// TIA Portal project "e045002v093" (V13)

(* hardware
DEVICE "S7-300 station_1"  S7-300 station
   slot 0: "Perfil soporte"  Rail  6ES7 390-1***0-0AA0
   slot 2: "U10.5"  CPU 313C  6ES7 313-5BG04-0AB0  V3.3
      slot 0: "Interfaz MPI_1"  MPI
      slot 2: "DI24/DO16_1"  DI24/DO16
      slot 3: "AI5/AO2_1"  AI5/AO2
      slot 4: "Contaje_1"  Counter
   slot 4: "U7.3"  CP 343-1 LEAN  6GK7 343-1CX10-0XE0  V3.0
   slot 5: "U13.5"  DI32xDC24V  6ES7 321-1BL00-0AA0
   slot 6: "U17.5"  DI32xDC24V  6ES7 321-1BL00-0AA0
   slot 7: "U21.5"  DI32 x 24VDC  6ES7 321-1BL00-0AA0
   slot 8: "U25.5"  DO16xRel. AC120V/230V  6ES7 322-1HH01-0AA0
   slot 9: "U27.5"  DO32xDC24V/0.5A  6ES7 322-1BL00-0AA0
   slot 10: "U35.5"  AO2 x 12bits  6ES7 332-5HB01-0AB0
DEVICE "U9.1"  KTP700 Basic PN
   slot 0: "HMI"  HMI  6AV2 123-2GB03-0AX0  13.0.1.0
   slot 1: "HMI_RT_1"  KTP700 Basic PN  6AV2 123-2GB03-0AX0  13.0.1.0
   slot 5: "U9.1.IE_CP_1"  Interfaz PROFINET
      slot 1: "Interfaz PROFINET_1"  Interfaz PROFINET
         slot 1: "Port_1"  Port
*)

// ===== PLC "U10.5"  CPU 313C =====
// protected blocks, not shown: "FB_CTR_MOT", "FC_MAQ_EST_16", "FC_MAQ_EST_32", "FC_PRC_ALA2", "fbSimContactor"

VAR_GLOBAL   // PLC tag table "00_Tabla de variables estándar"
   "CicIni" AT %M17.2 : Bool;
   "Clock_10.0_Hz" AT %M16.0 : Bool;
   "Clock_5.0_Hz" AT %M16.1 : Bool;
   "Clock_2.5_Hz" AT %M16.2 : Bool;
   "Clock_2.0_Hz" AT %M16.3 : Bool;
   "Clock_1.25_Hz" AT %M16.4 : Bool;
   "Clock_1.0_Hz" AT %M16.5 : Bool;
   "Clock_0.625_Hz" AT %M16.6 : Bool;
   "Clock_0.5_Hz" AT %M16.7 : Bool;
   "bit1" AT %M17.0 : Bool;
   "bit0" AT %M17.1 : Bool;
   "Rec_Todas" AT %M17.3 : Bool;
   "Tag_2" AT %M255.7 : Bool;
   "Tag_3" AT %M255.6 : Bool;
   "Tag_5" AT %M231.0 : Bool;
   "Tag_8" AT %T0 : Timer;
   "Ala_Nue" AT %M17.4 : Bool;
   "Ala_Pre" AT %M17.5 : Bool;
   "Sin_Ala" AT %M17.6 : Bool;
   "Contador" AT %MW18 : Word;
   "xpiSnsAscen_Aba_Par" AT %M248.2 : Bool;
   "_PeticiónPallet" AT %M251.5 : Bool;
   "Tag_9" AT %MB252 : Byte;
   "NoRstFilCompl" AT %M17.7 : Bool;   // No resetear "Fila Completa"
   "Set_TON_iSnsContadEmbal_1" AT %M232.0 : Bool;
   "Tag_4" AT %M241.1 : Bool;
   "Set_TON_iSnsContadEmbal_2" AT %M232.1 : Bool;
   "Set_TON_iSnsPerEmpCajAde" AT %M232.2 : Bool;
   "Cont_iSnsContadEmbal_1" AT %MW100 : Int;
   "Cont_iSnsContadEmbal_2" AT %MW102 : Int;
   "Cont_iSnsPerEmpCajAde" AT %MW104 : Int;
   "Cont_iSnsContadEmbal_3" AT %MW106 : Int;
   "Tag_6" AT %MD110 : Time;
   "Tag_7" AT %MD114 : Time;
   "Tag_10" AT %MD118 : Time;
   "Set_TON_iSnsContadEmbal_3" AT %M232.3 : Bool;
   "Tag_1" AT %T1 : Timer;
   "Tag_11" AT %M254.0 : Bool;
   "Tag_12" AT %M254.1 : Bool;
   "Tag_13" AT %M254.2 : Bool;
   "Tag_14" AT %M254.3 : Bool;
   "Tag_15" AT %M123.5 : Bool;
   "Tag_16" AT %M256.0 : Bool;
   "Tag_1200" AT %M255.0 : Bool;
   "Tag_17" AT %M255.1 : Bool;
   "Tag_18" AT %M33.5 : Bool;
   "Resum_ala_Fech" AT %M33.4 : Bool;
   "Hab_marcha1_2" AT %M50.7 : Bool;
   "T_espera_parada_21.26" AT %M50.5 : Bool;
   "MFRD" AT %M50.4 : Bool;
   "MIGS" AT %M50.6 : Bool;
   "i_SnsFinDosif" AT %I11.0 : Bool;   // Sensor final cinta dosificadora
END_VAR

VAR_GLOBAL   // PLC tag table "240_Memorias_Flancos"
   "xnHMI.Pls_Inc_Elem" AT %M240.0 : Bool;
   "xnHMI.Pls_Dec_Elem" AT %M240.1 : Bool;
   "xnHMI.Pls_Elem_Der" AT %M240.2 : Bool;
   "xnHMI.Pls_Elem_Izq" AT %M240.3 : Bool;
   "xnHMI.Pls_Inc_Fila" AT %M240.4 : Bool;
   "xnHMI.Pls_Dec_Fila" AT %M240.5 : Bool;
   "xnHMI.Pls_Fila_Sup" AT %M240.6 : Bool;
   "xnHMI.Pls_Fila_Inf" AT %M240.7 : Bool;
   "xpHMI.Pls_New_Fila" AT %M241.0 : Bool;
   "xpHMI.Pls_New_Elem" AT %M241.2 : Bool;
   "xpHMI.Pls_Kill_Elem" AT %M241.3 : Bool;
   "xnHMI.Pls_WR_Receta" AT %M241.4 : Bool;
   "xnHMI.Pls_RD_Receta" AT %M241.5 : Bool;
   "xpEditar_Recetas" AT %M241.6 : Bool;
   "xnHMI.Pls_Inc_Receta" AT %M241.7 : Bool;
   "xnHMI.Pls_Dec_Receta" AT %M242.0 : Bool;
   "xnHMI.Pls_Inc_Capa" AT %M242.1 : Bool;
   "xnHMI.Pls_Dec_Capa" AT %M242.2 : Bool;
   "xnHMI.Pls_Elem_+" AT %M242.3 : Bool;
   "xnHMI.Pls_Elem_-" AT %M242.4 : Bool;
   "xpHMI.Pls_CargarReceta" AT %M242.5 : Bool;
   "xpiPul_MarCiclo" AT %M242.6 : Bool;
   "xpiPul_HabTransp" AT %M242.7 : Bool;
   "xpiPul_HabDosif" AT %M243.0 : Bool;
   "xpiPul_HabCargPall" AT %M243.1 : Bool;
   "xpiPul_ResetAla" AT %M243.2 : Bool;
   "xpiSnsContadEmbal_1" AT %M243.3 : Bool;
   "xpiSnsContadEmbal_2" AT %M243.4 : Bool;
   "xniSnsContadEmbal_1" AT %M243.5 : Bool;
   "xniSnsContadEmbal_2" AT %M243.6 : Bool;
   "xpAUTO/MAN" AT %M243.7 : Bool;
   "xnAUTO/MAN" AT %M244.0 : Bool;
   "xniSnsPerEmpCajAde" AT %M244.1 : Bool;
   "xniSnsPallTrnsp_4" AT %M244.2 : Bool;
   "xniSnsPallTrnsp_5" AT %M244.3 : Bool;
   "xpiPul_MultiArr" AT %M244.4 : Bool;
   "xniPul_MultiArr" AT %M244.5 : Bool;
   "xpiPul_MultiAba" AT %M244.6 : Bool;
   "xniPul_MultiAba" AT %M244.7 : Bool;
   "xpiPul_MultiAde" AT %M245.0 : Bool;
   "xniPul_MultiAde" AT %M245.1 : Bool;
   "xpiPul_MultiAtr" AT %M245.2 : Bool;
   "xniPul_MultiAtr" AT %M245.3 : Bool;
   "xpiPul_Multi_A" AT %M245.4 : Bool;
   "xniPul_Multi_A" AT %M245.5 : Bool;
   "xpiPul_Multi_B" AT %M245.6 : Bool;
   "xniPul_Multi_B" AT %M245.7 : Bool;
   "xniSnsPlataf_Ade" AT %M246.0 : Bool;
   "xniSnsPlataf_Atr" AT %M246.1 : Bool;
   "xniSnsPallTrnsp_2" AT %M246.3 : Bool;
   "xpiSnsPallTrnsp_2" AT %M246.2 : Bool;
   "xpiSnsPallRetractil" AT %M246.4 : Bool;
   "xniSnsPallRetractil" AT %M246.5 : Bool;
   "xpiSnsPallTrnsp_4" AT %M246.6 : Bool;
   "xpiSnsPallTrnsp_5" AT %M246.7 : Bool;
   "xpiSnsEmpj_Ade_Par" AT %M247.0 : Bool;
   "xnPALLET_NO_FUERA_ASCENSOR" AT %M247.1 : Bool;
   "xpRECAMBIO_PALLET" AT %M247.2 : Bool;
   "xpiSnsPallEnAscen" AT %M247.3 : Bool;
   "xniSnsPallEnAscen" AT %M247.4 : Bool;
   "xpiSnsAltuPlata_Aba" AT %M247.5 : Bool;
   "xniSnsAltuPlata_Aba" AT %M247.6 : Bool;
   "xpiSnsAltuPlata_Arr" AT %M247.7 : Bool;
   "xniSnsAltuPlata_Arr" AT %M248.0 : Bool;
   "xpiSnsAscen_Arr" AT %M248.1 : Bool;
   "xnEditando_Recetas" AT %M248.3 : Bool;
   "xpHMI.Pls_RD_Receta" AT %M248.4 : Bool;
   "xp3s4" AT %M248.5 : Bool;
   "xp3s9" AT %M248.6 : Bool;
   "xpHMI.Pls_Inc_Figura_Sel" AT %M248.7 : Bool;
   "xpHMI.Pls_Inc_Capa_Editando" AT %M249.0 : Bool;
   "xpHMI.Pls_Dec_Capa_Editando" AT %M249.1 : Bool;
   "xpS_PriElemCapa" AT %M249.2 : Bool;
   "xnElemento_DESCARGADO" AT %M249.3 : Bool;
   "xpiSnsPerEmpCajAde" AT %M249.4 : Bool;
   "xpiSnsContadEmbal_3" AT %M249.5 : Bool;
   "xniSnsContadEmbal_3" AT %M249.6 : Bool;
END_VAR

VAR_GLOBAL   // PLC tag table "20_Recetas"
   "Editando_Recetas" AT %M20.0 : Bool;
   "RECETA_Editando" AT %MB21 : Byte;
   "CAPA_Editando" AT %MB22 : Byte;
END_VAR

VAR_GLOBAL   // PLC tag table "30_Proceso"
   "Elemento_CARGADO" AT %M30.0 : Bool;   // Avanzar en el dibujo
   "Nueva_CAPA" AT %M30.2 : Bool;   // Se terminó una capa
   "Elemento_DESCARGADO" AT %M30.1 : Bool;   // Retroceder en el dibujo
   "Nuevo_PALLET" AT %M30.3 : Bool;   // Se terminó un pallet
   "CICLO_Hab" AT %M30.4 : Bool;   // Máquina en ciclo automático
   "TRANSPORTES_Hab" AT %M30.5 : Bool;
   "DOSIFICADOR_Hab" AT %M30.6 : Bool;
   "CARGAPALLET_Hab" AT %M30.7 : Bool;
   "AUTO/MAN" AT %M31.0 : Bool;   // 1: AUTOMÁTICO / 0: MANUAL
   "ResumAla_Grave" AT %M31.1 : Bool;
   "ResumAla_General" AT %M31.2 : Bool;
   "ResumAla_TranspCaja_1" AT %M31.3 : Bool;
   "ResumAla_TranspCaja_2" AT %M31.4 : Bool;
   "ResumAla_Dosificador_1" AT %M31.5 : Bool;
   "ResumAla_Dosificador_2" AT %M31.6 : Bool;
   "ResumAla_CargaPallet_1" AT %M31.7 : Bool;
   "ResumAla_CargaPallet_2" AT %M32.0 : Bool;
   "ResumAla_CargaPallet_3" AT %M32.1 : Bool;
   "ResumAla_CargaPallet_4" AT %M32.2 : Bool;
   "ResumAla_TranspPall_1" AT %M32.3 : Bool;
   "ResumAla_TranspPall_2" AT %M32.4 : Bool;
   "ResumAla_Warnings" AT %M32.5 : Bool;
   "T_ResumAla_General" AT %M32.6 : Bool;
   "Esperando_Cajas" AT %M32.7 : Bool;
   "Cambio_Elemento" AT %M33.0 : Bool;
   "Elemento_DESCARGADO_scan" AT %M33.1 : Bool;
   "ResumAla_Dosificador_3" AT %M33.2 : Bool;
   "ResumAla_Dosificador_4" AT %M33.3 : Bool;
END_VAR

VAR_GLOBAL   // PLC tag table "Tabla I/O"
   "iPul_MultiArr" AT %E34.0 : Bool;   // Pulsador Multifunción Arriba
   "iPul_MultiAba" AT %E34.1 : Bool;   // Pulsador Multifunción Abajo
   "iPul_MultiAde" AT %E34.2 : Bool;   // Pulsador Multifunción Adelante
   "iPul_MultiAtr" AT %E34.3 : Bool;   // Pulsador Multifunción Atrás
   "iPul_Multi_A" AT %E34.4 : Bool;   // Pulsador Multifunción "A"
   "iPul_Multi_B" AT %E34.5 : Bool;   // Pulsador Multifunción "B"
   "iPul_ResetAla" AT %E34.6 : Bool;   // Pulsador Reset Alarmas
   "iiPul_Emerg" AT %E34.7 : Bool;   // Pulsador Parada de Emergencia en Pupitre
   "iPul_MarCiclo" AT %E32.0 : Bool;   // Pulsador Marcha de Ciclo
   "iiPul_ParaCiclo" AT %E32.1 : Bool;   // Pulsador Parada de Piclo
   "iPul_HabTransp" AT %E32.2 : Bool;   // Pulsador Habilitación Transporte de Entrada
   "iiPul_DeshTransp" AT %E32.3 : Bool;   // Pulsador Deshabilitación Transporte de Entrada
   "iPul_HabDosif" AT %E32.4 : Bool;   // Pulsador Habilitación Dosificador
   "iiPul_DeshDosif" AT %E32.5 : Bool;   // Pulsador Deshabilitación Dosificador
   "iPul_HabCargPall" AT %E32.6 : Bool;   // Pulsador Habilitación Carga de Pallet
   "iiPul_DeshCargPall" AT %E32.7 : Bool;   // Pulsador Deshabilitación Carga de Pallet
   "iSel_Auto/Man" AT %E33.0 : Bool;   // Selectora Automático/Manual
   "iiPul_EmergAlmac_1_AlmacManual" AT %E33.5 : Bool;   // Pulsador Operación Manual Almacén Pallets
   "iiPul_EmergAlmac_2" AT %E1.0 : Bool;   // Pulsador parada de emergencia en almacén
   "iPul_RstSegRetrAlmac" AT %E1.1 : Bool;   // Pulsador reset seguridades retractilador almacén
   "iiPul_EmergAscen" AT %E1.2 : Bool;   // Pulsador parada de emergencia en ascensor
   "iPul_RstSegRetrAscen" AT %E1.3 : Bool;   // Pulsador reset seguridades retractilador ascensor
   "iPul_RstSegRetrEntra" AT %E1.4 : Bool;   // Pulsador reset seguridades retractilador entrada
   "iPul_RstSegRetrSali" AT %E1.5 : Bool;   // Pulsador reset seguridades retractilador salida
   "iiPul_EmergMaq" AT %E1.6 : Bool;   // Pulsador parada de emergencia en máquina
   "iiPul_EmergTransp" AT %E1.7 : Bool;   // Pulsador parada de emergencia en transportes de alimentación
   "iVarEmpj_FLT" AT %E2.3 : Bool;   // Variador Empujador de Filas falla (FAULT)
   "iVarAscen_RDY" AT %E2.4 : Bool;   // Variador Ascensor listo (READY)
   "iVarAscen_FLT" AT %E2.5 : Bool;   // Variador Ascensor falla (FAULT)
   "iSnsEmpj_Atr_Par" AT %E3.1 : Bool;   // Sensor Empujador de Filas atrás parar
   "iSnsEmpj_Atr_Len" AT %E3.2 : Bool;   // Sensor Empujador de Filas atrás lento
   "iSnsEmpj_MedCamin" AT %E3.3 : Bool;   // Sensor Empujador de Filas a medio camino
   "iSnsEmpj_Ade_Len" AT %E3.4 : Bool;   // Sensor Empujador de Filas adelante lento
   "iSnsEmpj_Ade_Par" AT %E3.5 : Bool;   // Sensor Empujador de Filas adelante parar
   "iSnsEmpj_Abajo" AT %E3.6 : Bool;   // Sensor Empujador de Filas abajo
   "iSnsEmpj_Arriba" AT %E3.7 : Bool;   // Sensor Empujador de Filas arriba
   "iSnsSegTranspEntra" AT %E8.5 : Bool;   // Sensor Seguridad Transporte de entrada
   "iSnsSegEntraEmpj_1" AT %E8.6 : Bool;   // Sensor Seguridad Entrada Empujador de Filas 1
   "iSnsSegEntraEmpj_2" AT %E8.7 : Bool;   // Sensor Seguridad Entrada Empujador de Filas 2
   "iSnsSegAscen_1" AT %E9.2 : Bool;   // Sensor Seguridades acceso a Ascensor 1
   "iSnsSegAscen_2" AT %E9.3 : Bool;   // Sensor Seguridades acceso a Ascensor 2
   "iSnsSeg1Entra1Retrac" AT %E9.4 : Bool;   // Sensor Seguridades 1 Entrada 1 Retractilador
   "iSnsSeg2Entra1Retrac" AT %E9.5 : Bool;   // Sensor Seguridades 2 Entrada 1 Retractilador
   "iSnsSeg1Entra2Retrac" AT %E9.6 : Bool;   // Sensor Seguridades 1 Entrada 2 Retractilador
   "iSnsSeg2Entra2Retrac" AT %E9.7 : Bool;   // Sensor Seguridades 2 Entrada 2 Retractilador
   "iSeguridades" AT %E10.0 : Bool;   // Resumen de Seguridades
   "iTermMaq" AT %E10.1 : Bool;   // Resumen de térmicos en máquina
   "iTermTansp" AT %E10.2 : Bool;   // Resumen de térmicos en transportes
   "iSnsContadEmbal_3" AT %E10.4 : Bool;   // Sensor Contador de embalaje 3
   "oLuz_Segur" AT %A33.0 : Bool;   // Lámpara Seguridades
   "oLuz_CicloHab" AT %A33.1 : Bool;   // Lámpara Ciclo Habilitado
   "oLuz_TranspHab" AT %A33.2 : Bool;   // Lámpara Transportes de Alimentación Habilitados
   "oLuz_DosifHab" AT %A33.3 : Bool;   // Lámpara Dosificador Habilitado
   "oLuz_EmergMaq" AT %A33.5 : Bool;   // Lámpara Emergencia en Máquina
   "oLibre_A137" AT %A13.1 : Bool;
   "oResetVarEmpj" AT %A34.0 : Bool;   // Reset falla en variador Empujador de Filas
   "oResetVarDosif" AT %A34.2 : Bool;   // Reset falla en variador Dosificador
   "oEmpj_Subir" AT %A34.7 : Bool;
   "oLuz_ModoManual" AT %A16.6 : Bool;
   "oLuz_Baliza" AT %A16.7 : Bool;   // Baliza
   "oLibre_A175" AT %A17.5 : Bool;
   "oVal_Encolado" AT %A18.0 : Bool;   // Válvula de Encolado
   "oLuz_SegAscensor" AT %A19.4 : Bool;   // Lámpara Seguridades Ascensor
   "iwLibre_32.1" AT %EW524 : Word;
   "iwLibre_32.3" AT %EW526 : Word;
   "iwLibre_32.4" AT %EW528 : Word;
   "iwLibre_32.6" AT %EW530 : Word;
   "iwLibre_32.7" AT %EW532 : Word;
   "owVelRef_Dosif" AT %AW524 : Word;   // Velocidad de Referencia Variador Dosificador
   "owVelRef_Empuj" AT %AW526 : Word;   // Velocidad de Referencia Variador Empujador de Filas
   "owLibre_34.6" AT %AW514 : Word;
   "iVarEmpj_RDY" AT %E2.2 : Bool;   // Variador Empujador de Filas listo (READY)
   "oTranspPall2" AT %A13.3 : Bool;   // NO ESTÁ EN PLANOS - Marcha transporte de pallet 2 - Arrancador Suave -
   "oTranspPall3" AT %A13.4 : Bool;   // NO ESTÁ EN PLANOS - Marcha transporte de pallet 3 - Arrancador Suave -
   "iConf_Mar_Empu_Subir" AT %E33.1 : Bool;   // Confirmación K18: Empujador de Filas Subir
   "iConf_Mar_Empu_Bajar" AT %E33.2 : Bool;   // Confirmación K19: Empujador de Filas Bajar
   "iConf_Mar_Plataf_Adel" AT %E33.3 : Bool;   // Confirmación K21: Plataforma Carga Hacia Adelante
   "iConf_Mar_Plataf_Atra" AT %E33.4 : Bool;   // Confirmación K22: Plataforma Carga Hacia Atrás
END_VAR

VAR_GLOBAL   // PLC tag table "50_Transporte_Cajas"
   "MarTransp_21.10" AT %M50.0 : Bool;
   "MarTransp_21.22" AT %M50.1 : Bool;
   "MarTransp_21.24" AT %M50.2 : Bool;
   "MarTransp_21.26" AT %M50.3 : Bool;
   "iSnsCajaEn_21.22" AT %E7.0 : Bool;   // Sensor cajas acumuladas en transporte 21.22
   "iSnsCajaEn_21.26" AT %E7.1 : Bool;   // Sensor cajas acumuladas en transporte 21.26
   "oTransp_21.10" AT %A12.0 : Bool;   // Marcha cinta 21.10 del transporte de Alimentación - K4 -
   "oTransp_21.22" AT %A12.1 : Bool;   // Marcha rolos 21.22 del transporte de Alimentación - K6 -
   "oTransp_21.24" AT %A12.2 : Bool;   // Marcha cinta 21.24 del transporte de Alimentación - K8 -
   "oTransp_21.26" AT %A12.3 : Bool;   // Marcha rolos 21.26 del transporte de Alimentación - K10 -
END_VAR

VAR_GLOBAL   // PLC tag table "230_Alarmas"
   "Falla_CARGAPALLET" AT %M230.3 : Bool;
   "Color_Alarmas" AT %MB231 : Byte;
   "Habil_Ala_82" AT %M230.4 : Bool;   // Habilita la activación de la alarma de Barrera a la salida de la Envolvedora
END_VAR

VAR_GLOBAL   // PLC tag table "60_Dosificador"
   "MarBandaDosif" AT %M60.0 : Bool;
   "MarTranspEntra1" AT %M60.1 : Bool;
   "MarTranspEntra2" AT %M60.5 : Bool;
   "Act_GiraCaja" AT %M60.2 : Bool;
   "Act_EmpujaCaja" AT %M60.3 : Bool;
   "Act_StopCaja" AT %M60.4 : Bool;
   "iVarDosif_RDY" AT %E2.6 : Bool;   // Variador Cinta Dosificadora listo (READY)
   "iVarDosif_FLT" AT %E2.7 : Bool;   // Variador Cinta Dosificadora falla (FAULT)
   "iSnsEmpCaja_Ade" AT %E3.0 : Bool;   // Sensor Empujador de Cajas adelante
   "iSnsSolapaAbierta" AT %E7.2 : Bool;   // Sensor solapa abierta
   "iSnsPerEmpCajAde" AT %E7.3 : Bool;   // Sensor permiso Empujador de Cajas adelante
   "iSnsContadEmbal_1" AT %E8.3 : Bool;   // Sensor Contador de embalaje 1
   "iSnsContadEmbal_2" AT %E8.4 : Bool;   // Sensor Contador de embalaje 2
   "oTransp_Entra1" AT %A12.4 : Bool;   // Marcha rolos transporte de entrada 1 - K14 -
   "oTransp_Entra2" AT %A12.5 : Bool;   // Marcha rolos transporte de entrada 2 - K15 -
   "oEmpj_Subir_old" AT %A12.6 : Bool;   // Marcha Empujador de Filas subir - K18 -
   "oEmpj_Bajar" AT %A12.7 : Bool;   // Marcha Empujador de Filas bajar - K19 -
   "oEmpjFrenoAvaRet" AT %A16.0 : Bool;   // Liberar Freno del Empujador de Filas - Avance/Retroceso - K27.1 -
   "oEmpjFrenoSubBaj" AT %A16.1 : Bool;   // Liberar Freno del Empujador de Filas - Subir/Bajar - K27.2 -
   "oMarBanDosif" AT %A17.0 : Bool;   // Marcha Banda Dosificadora - V1 -
   "oMarEmpj" AT %A17.1 : Bool;   // Marcha Empujador de Filas - V2 -
   "oInvGiroEmpj" AT %A17.2 : Bool;   // Invertir giro marcha Empujador de Filas - V2 -
   "oVal_GiraCaja" AT %A18.1 : Bool;   // Válvula de Girador de Cajas
   "oVal_EmpujaCaja" AT %A18.2 : Bool;   // Válvula de Empujador de Cajas
   "oVal_StopCaja" AT %A18.3 : Bool;   // Válvula de Stop de Cajas
   "Dosif_SPVel" AT %MD62 : Real;
   "Levantar_Stop_Aux" AT %M60.6 : Bool;
   "Terminar_Empujador_Aux" AT %M60.7 : Bool;
   "mem_Terminar_Empujador_Aux" AT %M61.0 : Bool;
   "_Cx_Temp" AT %M61.1 : Bool;
   "Titilar_Dosificador" AT %M61.2 : Bool;
   "_Caja_en_Medio" AT %M61.3 : Bool;   // Prueba
   "Frena_Dosif" AT %M61.4 : Bool;
   "Anterior_Vertical" AT %M61.5 : Bool;
   "Detener_Dosificador" AT %M61.6 : Bool;
   "Scan_iSnsContadEmbal_1" AT %M61.7 : Bool;
END_VAR

VAR_GLOBAL   // PLC tag table "200_Máq_Estados"
   "_c1" AT %M200.0 : Bool;   // Ir a Estado 1
   "_c2" AT %M200.1 : Bool;   // Ir a Estado 2
   "_c3" AT %M200.2 : Bool;   // Ir a Estado 3
   "_c4" AT %M200.3 : Bool;   // Ir a Estado 4
   "_c5" AT %M200.4 : Bool;   // Ir a Estado 5
   "_c6" AT %M200.5 : Bool;   // Ir a Estado 6
   "_c7" AT %M200.6 : Bool;   // Ir a Estado 7
   "_c8" AT %M200.7 : Bool;   // Ir a Estado 8
   "_c9" AT %M201.0 : Bool;   // Ir a Estado 9
   "_c10" AT %M201.1 : Bool;   // Ir a Estado 10
   "_c11" AT %M201.2 : Bool;   // Ir a Estado 11
   "_c12" AT %M201.3 : Bool;   // Ir a Estado 12
   "_c13" AT %M201.4 : Bool;   // Ir a Estado 13
   "_c14" AT %M201.5 : Bool;   // Ir a Estado 14
   "_c15" AT %M201.6 : Bool;   // Ir a Estado 15
   "_c16" AT %M201.7 : Bool;   // Ir a Estado 16
   "_c17" AT %M202.0 : Bool;   // Ir a Estado 17
   "_c18" AT %M202.1 : Bool;   // Ir a Estado 18
   "_c19" AT %M202.2 : Bool;   // Ir a Estado 19
   "_c20" AT %M202.3 : Bool;   // Ir a Estado 20
   "_c21" AT %M202.4 : Bool;   // Ir a Estado 21
   "_c22" AT %M202.5 : Bool;   // Ir a Estado 22
   "_c23" AT %M202.6 : Bool;   // Ir a Estado 23
   "_c24" AT %M202.7 : Bool;   // Ir a Estado 24
   "_c25" AT %M203.0 : Bool;   // Ir a Estado 25
   "_c26" AT %M203.1 : Bool;   // Ir a Estado 26
   "_c27" AT %M203.2 : Bool;   // Ir a Estado 27
   "_c28" AT %M203.3 : Bool;   // Ir a Estado 28
   "_c29" AT %M203.4 : Bool;   // Ir a Estado 29
   "_c30" AT %M203.5 : Bool;   // Ir a Estado 30
   "_c31" AT %M203.6 : Bool;   // Ir a Estado 31
   "_c32" AT %M203.7 : Bool;   // Ir a Estado 32
   "_p1" AT %M204.0 : Bool;   // Forzar Estado 1
   "_p2" AT %M204.1 : Bool;   // Forzar Estado 2
   "_p3" AT %M204.2 : Bool;   // Forzar Estado 3
   "_p4" AT %M204.3 : Bool;   // Forzar Estado 4
   "_p5" AT %M204.4 : Bool;   // Forzar Estado 5
   "_p6" AT %M204.5 : Bool;   // Forzar Estado 6
   "_p7" AT %M204.6 : Bool;   // Forzar Estado 7
   "_p8" AT %M204.7 : Bool;   // Forzar Estado 8
   "_p9" AT %M205.0 : Bool;   // Forzar Estado 9
   "_p10" AT %M205.1 : Bool;   // Forzar Estado 10
   "_p11" AT %M205.2 : Bool;   // Forzar Estado 11
   "_p12" AT %M205.3 : Bool;   // Forzar Estado 12
   "_p13" AT %M205.4 : Bool;   // Forzar Estado 13
   "_p14" AT %M205.5 : Bool;   // Forzar Estado 14
   "_p15" AT %M205.6 : Bool;   // Forzar Estado 15
   "_p16" AT %M205.7 : Bool;   // Forzar Estado 16
   "_p17" AT %M206.0 : Bool;   // Forzar Estado 17
   "_p18" AT %M206.1 : Bool;   // Forzar Estado 18
   "_p19" AT %M206.2 : Bool;   // Forzar Estado 19
   "_p20" AT %M206.3 : Bool;   // Forzar Estado 20
   "_p21" AT %M206.4 : Bool;   // Forzar Estado 21
   "_p22" AT %M206.5 : Bool;   // Forzar Estado 22
   "_p23" AT %M206.6 : Bool;   // Forzar Estado 23
   "_p24" AT %M206.7 : Bool;   // Forzar Estado 24
   "_p25" AT %M207.0 : Bool;   // Forzar Estado 25
   "_p26" AT %M207.1 : Bool;   // Forzar Estado 26
   "_p27" AT %M207.2 : Bool;   // Forzar Estado 27
   "_p28" AT %M207.3 : Bool;   // Forzar Estado 28
   "_p29" AT %M207.4 : Bool;   // Forzar Estado 29
   "_p30" AT %M207.5 : Bool;   // Forzar Estado 30
   "_p31" AT %M207.6 : Bool;   // Forzar Estado 31
   "_p32" AT %M207.7 : Bool;   // Forzar Estado 32
   "1s1" AT %M208.0 : Bool;   // DOSIFICADOR 1: REPOSO
   "1s2" AT %M208.1 : Bool;   // DOSIFICADOR 2: METE CAJA
   "1s3" AT %M208.2 : Bool;   // DOSIFICADOR 3: FIGURA H
   "1s4" AT %M208.3 : Bool;   // DOSIFICADOR 4: FIGURA V
   "1s5" AT %M208.4 : Bool;   // DOSIFICADOR 5: FIGURA HH
   "1s6" AT %M208.5 : Bool;   // DOSIFICADOR 6: ALMACENA CAJA
   "1s7" AT %M208.6 : Bool;   // DOSIFICADOR 7: ALMACENA CAJA
   "1s8" AT %M208.7 : Bool;   // DOSIFICADOR 8: METE CAJA
   "1s9" AT %M209.0 : Bool;   // DOSIFICADOR 9: ALMACENA CAJA
   "1s10" AT %M209.1 : Bool;   // DOSIFICADOR 10: ACOMODO
   "1s11" AT %M209.2 : Bool;   // DOSIFICADOR 11: EMPUJA
   "1s12" AT %M209.3 : Bool;   // DOSIFICADOR 12: ESPERA
   "1s13" AT %M209.4 : Bool;   // DOSIFICADOR 13: ALMACENA CAJA
   "1s14" AT %M209.5 : Bool;   // DOSIFICADOR 14: METIENDO H
   "1s15" AT %M209.6 : Bool;   // DOSIFICADOR 15: METIENDO V
   "1s16" AT %M209.7 : Bool;   // DOSIFICADOR 16: METIENDO HH
   "1s17" AT %M210.0 : Bool;
   "1s18" AT %M210.1 : Bool;
   "1s19" AT %M210.2 : Bool;
   "1s20" AT %M210.3 : Bool;
   "1s21" AT %M210.4 : Bool;
   "1s22" AT %M210.5 : Bool;
   "1s23" AT %M210.6 : Bool;
   "1s24" AT %M210.7 : Bool;
   "1s25" AT %M211.0 : Bool;
   "1s26" AT %M211.1 : Bool;
   "1s27" AT %M211.2 : Bool;
   "1s28" AT %M211.3 : Bool;
   "1s29" AT %M211.4 : Bool;
   "1s30" AT %M211.5 : Bool;
   "1s31" AT %M211.6 : Bool;
   "1s32" AT %M211.7 : Bool;
   "2s1" AT %M212.0 : Bool;   // CARGA_PALLET 1: REPOSO
   "2s2" AT %M212.1 : Bool;   // CARGA_PALLET 2: PLATAFORMA CARGADA
   "2s3" AT %M212.2 : Bool;   // CARGA_PALLET 3: SUBIR RÁPIDO
   "2s4" AT %M212.3 : Bool;   // CARGA_PALLET 4: SUBIR LENTO
   "2s5" AT %M212.4 : Bool;   // CARGA_PALLET 5: ADELANTAR
   "2s6" AT %M212.5 : Bool;   // CARGA_PALLET 6: PONER MORDAZAS
   "2s7" AT %M212.6 : Bool;   // CARGA_PALLET 7: PONER BRAZO
   "2s8" AT %M212.7 : Bool;   // CARGA_PALLET 8: RETIRAR
   "2s9" AT %M213.0 : Bool;   // CARGA_PALLET 9: LIBERAR
   "2s10" AT %M213.1 : Bool;   // CARGA_PALLET 10: SACAR BRAZO
   "2s11" AT %M213.2 : Bool;   // CARGA_PALLET 11: IR ZONA SUPERIOR LENTO
   "2s12" AT %M213.3 : Bool;   // CARGA_PALLET 12: RECAMBIO PALLET
   "2s13" AT %M213.4 : Bool;   // CARGA_PALLET 13: IR ZONA INFERIOR RÁPIDO
   "2s14" AT %M213.5 : Bool;   // CARGA_PALLET 14: IR ZONA INFERIOR LENTO
   "2s15" AT %M213.6 : Bool;   // CARGA_PALLET 15: METER PISTÓN
   "2s16" AT %M213.7 : Bool;   // CARGA_PALLET 16: SACAR PISTÓN
   "2s17" AT %M214.0 : Bool;   // CARGA_PALLET 17: SUBIR LENTO
   "2s18" AT %M214.1 : Bool;
   "2s19" AT %M214.2 : Bool;
   "2s20" AT %M214.3 : Bool;
   "2s21" AT %M214.4 : Bool;
   "2s22" AT %M214.5 : Bool;
   "2s23" AT %M214.6 : Bool;
   "2s24" AT %M214.7 : Bool;
   "2s25" AT %M215.0 : Bool;
   "2s26" AT %M215.1 : Bool;
   "2s27" AT %M215.2 : Bool;
   "2s28" AT %M215.3 : Bool;
   "2s29" AT %M215.4 : Bool;
   "2s30" AT %M215.5 : Bool;
   "2s31" AT %M215.6 : Bool;
   "2s32" AT %M215.7 : Bool;
   "dc_" AT %MD200 : DWord;   // Concatenadora
   "dp_" AT %MD204 : DWord;   // Prioritaria
   "ds1" AT %MD208 : DWord;   // Estado del DOSIFICADOR
   "ds2" AT %MD212 : DWord;   // Estado de la PLATAFORMA
   "ErrForz_1" AT %M220.0 : Bool;
   "ErrTrans_1" AT %M220.1 : Bool;
   "ErrForz_2" AT %M220.2 : Bool;
   "ErrTrans_2" AT %M220.3 : Bool;
   "ws3" AT %MW216 : Word;   // Estado del EMPUJADOR
   "ErrForz_3" AT %M220.4 : Bool;
   "ErrTrans_3" AT %M220.5 : Bool;
   "3s1" AT %M216.0 : Bool;   // EMPUJADOR 1: REPOSO
   "3s2" AT %M216.1 : Bool;   // EMPUJADOR 2: ADELANTAR MEDIO
   "3s3" AT %M216.2 : Bool;   // EMPUJADOR 3: SUBIR
   "3s4" AT %M216.3 : Bool;   // EMPUJADOR 4: RETROCERDER RÁPIDO
   "3s5" AT %M216.4 : Bool;   // EMPUJADOR 5: RETROCERDER LENTO
   "3s6" AT %M216.5 : Bool;   // EMPUJADOR 6: BAJAR
   "3s7" AT %M216.6 : Bool;   // EMPUJADOR 7: ESPERA PLATAFORMA
   "3s8" AT %M216.7 : Bool;   // EMPUJADOR 8: ADELANTAR FINAL
   "3s9" AT %M217.0 : Bool;   // EMPUJADOR 9: ADELANTAR FINAL y HAB FILA
   "3s10" AT %M217.1 : Bool;   // EMPUJADOR 10: ADELANTAR LENTO FINAL
   "3s11" AT %M217.2 : Bool;
   "3s12" AT %M217.3 : Bool;
   "3s13" AT %M217.4 : Bool;
   "3s14" AT %M217.5 : Bool;
   "3s15" AT %M217.6 : Bool;
   "3s16" AT %M217.7 : Bool;
   "wc_" AT %MW200 : Word;   // Concatenadora
   "wp_" AT %MW204 : Word;   // Prioritaria
   "ErrForz_4" AT %M220.6 : Bool;
   "ErrTrans_4" AT %M220.7 : Bool;
   "ws4" AT %MW218 : Word;
   "4s1" AT %M218.0 : Bool;   // ELEMENTO_HH 1: REPOSO
   "4s2" AT %M218.1 : Bool;   // ELEMENTO_HH 2: ESPERA CAJA 2
   "4s3" AT %M218.2 : Bool;   // ELEMENTO_HH 3: FRENANDO CAJA 2
   "4s4" AT %M218.3 : Bool;   // ELEMENTO_HH 4: ALMACENA CAJAS
   "4s5" AT %M218.4 : Bool;
   "4s6" AT %M218.5 : Bool;
   "4s7" AT %M218.6 : Bool;
   "4s8" AT %M218.7 : Bool;
   "4s9" AT %M219.0 : Bool;
   "4s10" AT %M219.1 : Bool;
   "4s11" AT %M219.2 : Bool;
   "4s12" AT %M219.3 : Bool;
   "4s13" AT %M219.4 : Bool;
   "4s14" AT %M219.5 : Bool;
   "4s15" AT %M219.6 : Bool;
   "4s16" AT %M219.7 : Bool;
END_VAR

VAR_GLOBAL   // PLC tag table "70_Empujador"
   "Empujador_MEDIO" AT %M70.0 : Bool;
   "Empujador_ADE_PARAR" AT %M70.1 : Bool;
   "Empujador_ARR" AT %M70.2 : Bool;
   "Empujador_ATR_LENTO" AT %M70.3 : Bool;
   "Empujador_ATR_PARAR" AT %M70.4 : Bool;
   "Empujador_ADE_LENTO" AT %M70.5 : Bool;
   "Empujador_ABA" AT %M70.6 : Bool;
   "E_Plataforma_en_Posición" AT %M70.7 : Bool;
   "E_Elemento_Cargado" AT %M71.0 : Bool;
   "S_ÚltElemFila" AT %M71.1 : Bool;   // Indica que el elemento seleccionado es el último de una fila
   "S_ÚltFilCapa" AT %M71.2 : Bool;
   "PEDIDO_de_CAJA" AT %M71.3 : Bool;
   "Espacio_Mesa_Intermedia" AT %M71.4 : Bool;
   "Fila_Completa" AT %M71.5 : Bool;
   "Ord_Empujad_Subir" AT %M71.6 : Bool;
   "Ord_Empujad_Bajar" AT %M71.7 : Bool;
   "Empuj_FrenoSubBajLibre" AT %M72.0 : Bool;
   "Ord_Empujad_Adel" AT %M72.1 : Bool;
   "Ord_Empujad_Atr" AT %M72.2 : Bool;
   "Empuj_SPVel_AdeAtr" AT %MD74 : Real;
   "EMPUJ_MED_CAM" AT %M72.3 : Bool;
   "_Último_Elemento_Temp" AT %M72.4 : Bool;   // BORRAR
   "_Temp" AT %M72.5 : Bool;   // BORRAR
   "Posición_Empujador_Ade-Atr" AT %MB73 : Byte;
   "EmpujaFil_Buscar_AtrParar" AT %M72.6 : Bool;
   "EmpujaFil_Buscar_AtrLento" AT %M72.7 : Bool;
   "EmpujaFil_Buscar_MedioCam" AT %M78.0 : Bool;
   "EmpujaFil_Buscar_AdeLento" AT %M78.1 : Bool;
   "EmpujaFil_Buscar_AdeParar" AT %M78.2 : Bool;
   "PosAnt_Empujador_Ade-Atr" AT %MB79 : Byte;
   "S_PriElemCapa" AT %M78.3 : Bool;
   "Medio_Camino" AT %M78.4 : Bool;
END_VAR

VAR_GLOBAL   // PLC tag table "80_Carga_Pallets"
   "iSnsPlataf_Atr" AT %E4.0 : Bool;   // Sensor Plataforma de Carga atrás
   "iSnsPlataf_Ade" AT %E4.1 : Bool;   // Sensor Plataforma de Carga adelante
   "iSnsRetEmpuBrazo" AT %E4.2 : Bool;   // Sensor Empujador en Brazo retirar (Plataforma Pos. Intermedia)
   "iSnsAscen_Aba_Par" AT %E4.3 : Bool;   // Sensor Ascensor abajo parar
   "iSnsAscen_Aba_Len" AT %E4.4 : Bool;   // Sensor Ascensor abajo lento
   "iSnsUltCapForm_2" AT %E4.5 : Bool;   // Sensor Última Capa de Formato _2
   "iSnsUltCapForm_1" AT %E4.6 : Bool;   // Sensor Última Capa de Formato _1
   "iSnsAscen_Arr" AT %E4.7 : Bool;   // Sensor Ascensor arriba
   "iSnsCerrSegAscen" AT %E5.0 : Bool;   // Sensor Cerrojo de Seguridad del ascensor
   "iSnsTopLat_Izq" AT %E6.0 : Bool;   // Sensor Tope Lateral Izquierdo
   "iSnsTopLat_Der" AT %E6.1 : Bool;   // Sensor Tope Lateral Derecho
   "iSnsTopPlat_Atr" AT %E6.2 : Bool;   // Sensor Tope Plataforma atrás
   "iSnsBarrDesc_Atr" AT %E6.3 : Bool;   // Sensor Pistón en Barra de Descarga atrás
   "iifcSegCadenas" AT %E6.4 : Bool;   // Finales de carrera Seguridades Cadena
   "ifcSegAscen_Arr" AT %E6.5 : Bool;   // Final de carrera Seguridad Ascensor arriba
   "iSnsCapFormPlat" AT %E7.4 : Bool;   // Sensor Capa formada en pallet
   "iSnsAltuPlata_Arr" AT %E7.5 : Bool;   // Sensor altura Plataforma arriba
   "iSnsAltuPlata_Aba" AT %E7.6 : Bool;   // Sensor altura Plataforma abajo
   "iSnsSegAscenBajar" AT %E8.1 : Bool;   // Sensor Seguridad Ascensor bajar
   "oPlataCarg_Ade" AT %A13.0 : Bool;   // Marcha Plataforma de Carga hacia adelante - K21 -
   "oPlataCarg_Atr" AT %A13.7 : Bool;   // Marcha Plataforma de Carga hacia atrás - K22 -
   "oPlataCargFreno" AT %A16.2 : Bool;   // Liberar Freno de la Plataforma de Carga - K27.3 -
   "oVal_BrazoDescar" AT %A18.4 : Bool;   // Válvula de Brazo de Descarga
   "oVal_EmpujBrazo" AT %A18.5 : Bool;   // Válvula de Empujador en Brazo de Descarga
   "oVal_MordazaFin" AT %A18.6 : Bool;   // Válvula de Mordaza Final
   "oVal_MordazasLat" AT %A18.7 : Bool;   // Válvula de Mordazas Laterales
   "Orden_Descargar" AT %M84.0 : Bool;
   "Poner_Mordazas" AT %M84.1 : Bool;
   "Ascensor_Subir_Lento" AT %M84.2 : Bool;
   "Ascensor_Posicionado" AT %M84.3 : Bool;
   "Plataforma_Adelante" AT %M84.4 : Bool;
   "Mordazas_Puestas" AT %M84.5 : Bool;
   "Brazo_Puesto" AT %M84.6 : Bool;
   "Plataforma_Atrás" AT %M84.7 : Bool;
   "Pistón_en_Brazo_Atrás" AT %M85.0 : Bool;
   "Brazo_y_Mordazas_Fuera" AT %M85.1 : Bool;
   "Última_Capa" AT %M85.2 : Bool;
   "Ascensor_Zona_Superior" AT %M85.3 : Bool;
   "PALLET_LLENO_SE_FUE" AT %M85.4 : Bool;
   "Ascensor_Casi_Zona_Inf" AT %M85.5 : Bool;
   "Ascensor_Zona_Inferior" AT %M85.6 : Bool;
   "Capa_en_Plataforma" AT %M85.7 : Bool;
   "Plataforma_FrenoLibre" AT %M86.0 : Bool;
   "Ord_Plataforma_Ade" AT %M86.1 : Bool;
   "Ord_Plataforma_Atr" AT %M86.2 : Bool;
   "oMarAscen" AT %A17.3 : Bool;   // Marcha Ascensor - V3 -
   "oInvGiroAscen" AT %A17.4 : Bool;   // Invertir giro marcha Ascensor - V3 -
   "oResetVarAscen" AT %A34.1 : Bool;   // Reset falla en variador Ascensor
   "owVelRef_Ascen" AT %AW512 : Word;   // Velocidad de Referencia Variador Ascensor
   "Ord_Ascensor_Subir" AT %M86.3 : Bool;
   "Ord_Ascensor_Bajar" AT %M86.4 : Bool;
   "Ord_Valv_Brazo" AT %M86.5 : Bool;
   "Ord_Valv_Pistón_Brazo" AT %M86.6 : Bool;
   "Ord_Mordazas" AT %M86.7 : Bool;
   "Vel_Ref_Ascensor" AT %MD80 : Real;
   "Petición_Plataforma_Ade" AT %M87.0 : Bool;
   "Petición_Plataforma_Atr" AT %M87.1 : Bool;
   "Poner_Pistón" AT %M87.2 : Bool;
   "Mem_Pistón" AT %M87.3 : Bool;
   "PosiciónPlataf_Ade-Atr" AT %MB88 : Byte;
   "PosiciónPlataf_Arr-Aba" AT %MB89 : Byte;
   "Brazo_Descarga_Man" AT %M87.4 : Bool;
END_VAR

VAR_GLOBAL   // PLC tag table "90_Transporte_Pallets"
   "iSnsPallTrnsp_2" AT %E5.1 : Bool;   // Sensor Pallet en Transporte 2
   "iSnsPallTrnsp_4" AT %E5.2 : Bool;   // Sensor Pallet en Transporte 4
   "iSnsPallTrnsp_5" AT %E5.3 : Bool;   // Sensor Pallet en Transporte 5
   "iSnsPallDescar" AT %E5.4 : Bool;   // Sensor Pallet en Descarga
   "iSnsAlmacPall_Arr" AT %E5.5 : Bool;   // Sensor Almacén de Pallets arriba
   "iSnsAlmacPall_Aba" AT %E5.7 : Bool;   // Sensor Almacén de Pallets abajo
   "iSnsPallEnAlmac" AT %E7.7 : Bool;   // Sensor de pallet en Almacén
   "iSnsPallEnAscen" AT %E8.0 : Bool;   // Sensor de pallet en Ascensor
   "iSnsPallRetractil" AT %E8.2 : Bool;   // Sensor pallet en Retractiladora
   "iSnsSegAlmac_1" AT %E9.0 : Bool;   // Sensor Seguridades Almacén 1
   "iSnsSegAlmac_2" AT %E9.1 : Bool;   // Sensor Seguridades Almacén 2
   "iPul_SubirAlmac" AT %E33.6 : Bool;   // Pulsador levantar almacén pallet
   "iPul_DedosAlmac" AT %E33.7 : Bool;   // Pulsador "dedos" almacén pallet
   "oTranspPall1" AT %A13.2 : Bool;   // Marcha transporte de pallet 1 - Arrancador Suave -
   "oTranspPall4" AT %A13.5 : Bool;   // Marcha transporte de pallet 4 - Arrancador Suave -
   "oTranspPall5" AT %A13.6 : Bool;   // Marcha transporte de pallet 5 - Arrancador Suave -
   "oVlvTulipaArrastre" AT %A16.5 : Bool;   // Válvula de Tulipa de arrastre
   "oVal_AlmacPallet" AT %A19.0 : Bool;   // Válvula de Almacén de Pallets
   "oVal_DedosAlmPall" AT %A19.1 : Bool;   // Válvula de Dedos en Almacén de Pallets
   "oVal_StopPallet" AT %A19.2 : Bool;   // Válvula de Stop de Pallets
   "oLuz_SegAmacPall" AT %A19.3 : Bool;   // Lámpara Seguridades Almacén
   "oLuz_SegRetrac1" AT %A19.5 : Bool;   // Lámpara Seguridades Retractilador 1
   "oLuz_SegRetrac2" AT %A19.6 : Bool;   // Lámpara Seguridades Retractilador 2
   "oLuz_SegTransPallet" AT %A19.7 : Bool;   // Lámpara Seguridades Transporte de Pallets
   "oLuz_CargPallHab" AT %A33.4 : Bool;   // Lámpara Carga de Pallet Habilitada
   "oLuz_EmergAlmac" AT %A33.6 : Bool;   // Lámpara Emergencia en Almacén de Pallets
   "oTranspPall3Freno" AT %A16.4 : Bool;   // Liberar Freno del transporte de pallet 3 - K27.5 -
   "OrdMar_TranspPall_1" AT %M90.0 : Bool;
   "OrdMar_TranspPall_2" AT %M90.1 : Bool;
   "OrdMar_TranspPall_3" AT %M90.2 : Bool;
   "OrdMar_TranspPall_4" AT %M90.3 : Bool;
   "OrdMar_TranspPall_5" AT %M90.4 : Bool;
   "TranspPall3_FrenoLibre" AT %M90.5 : Bool;
   "OrdVal_AlmacPall" AT %M90.6 : Bool;
   "OrdVal_DedosAlmac" AT %M90.7 : Bool;
   "DEDOS_ABIERTOS" AT %M91.0 : Bool;
   "ALMACÉN_Hab" AT %M91.1 : Bool;
   "BuscaPallet_Realizada" AT %M91.2 : Bool;
   "TranspPall_1_Detenido" AT %M91.3 : Bool;
   "Tonof_PALLET_EN_ASCENSOR" AT %M91.4 : Bool;
   "STOP_PALLET_ABIERTO" AT %M91.5 : Bool;
   "OrdVal_StopPallet" AT %M91.6 : Bool;
   "RECAMBIO_PALLET" AT %M91.7 : Bool;
   "PALLET_PARA_ASCENSOR" AT %M92.0 : Bool;
   "PALLET_NO_FUERA_ASCENSOR" AT %M92.1 : Bool;
   "TRANSP_2_POR_RECAMBIO" AT %M92.2 : Bool;
   "TRANSP_2_POR_ENVÍO" AT %M92.3 : Bool;
   "PALLET_SALIO_TRANSP_2" AT %M92.4 : Bool;
   "ZONA_ENVOLVEDORA_LIBRE" AT %M92.5 : Bool;
   "PALLET_EN_ENVOLVEDORA" AT %M92.6 : Bool;
   "ZONA_ETIQUETADORA_LIBRE" AT %M92.7 : Bool;
   "PALLET_EN_ETIQUETADORA" AT %M93.0 : Bool;
   "PALLET_FUERA_TRANSP_5" AT %M93.1 : Bool;
   "PALLET_DENTRO_TRANSP_5" AT %M93.2 : Bool;
   "TRANSP_3_POR_PEDIDO" AT %M93.3 : Bool;
   "TRANSP_3_POR_ENVÍO" AT %M93.4 : Bool;
   "TRANSP_4_POR_PEDIDO" AT %M93.5 : Bool;
   "TRANSP_4_POR_ENVÍO" AT %M93.6 : Bool;
   "TRANSP_5_POR_PEDIDO" AT %M93.7 : Bool;
   "PALLET_EN_ZONA_DESCARGA" AT %M94.0 : Bool;
   "ZONA_DESCARGA_LIBRE" AT %M94.1 : Bool;
   "PERMISO_ASCENSOR_BAJAR" AT %M94.2 : Bool;
   "TRANSP_1_POR_ENVÍO" AT %M94.3 : Bool;
   "TRANSP_1_POR_NUEVO_PALLET" AT %M94.4 : Bool;
   "TRANSP_1_POR_RECAMBIO" AT %M94.5 : Bool;
   "TRANSP_5_POR_ENVÍO" AT %M94.6 : Bool;
   "HAY_QUE_RECAMBIAR" AT %M94.7 : Bool;
   "TRANSP_2_VACÍO" AT %M95.0 : Bool;
   "PEDIDO_PALLET_ASCENSOR_con_pallet" AT %M95.1 : Bool;
   "PALLET_EN_ALMACEN" AT %M95.2 : Bool;
   "PEDIDO_PALLET_ASCENSOR_sin_pallet" AT %M95.3 : Bool;
   "PALLET_EN_ASCENSOR" AT %M95.4 : Bool;
   "Pallet_Envolvedora_a_Etiquetadora" AT %M95.5 : Bool;
   "Pallet_Etiquetadora_a_Transporte5" AT %M95.6 : Bool;
   "Pallet_Transporte5_a_Descarga" AT %M95.7 : Bool;
   "Pallet_Transporte2_a_Envolvedora" AT %M96.0 : Bool;
   "Pallet_Transporte1_a_Transporte2" AT %M96.1 : Bool;
   "Nueva_Etiqueta" AT %M96.2 : Bool;
   "iSnsAlmacPall_Med" AT %E5.6 : Bool;   // Sensor Almacén de Pallets medio
   "Posición_Almacén" AT %MB97 : Byte;
   "STOP_PALLET_ON" AT %M96.3 : Bool;
   "Pre-OrdMar_TranspPall_3" AT %M96.4 : Bool;
END_VAR

VAR_GLOBAL   // PLC tag table "I/O Intercambio Etiquetadora"
   "iHome_Pistón" AT %E10.3 : Bool;   // Home Pistón KETAN
   "iFin_Ciclo_Ketan" AT %E6.7 : Bool;   // Pallet etiquetado OK ó BYPASS
   "oEtiquetar_Pallet" AT %A33.7 : Bool;   // Pallet en transporte 4 para etiquetar
END_VAR

VAR_GLOBAL   // PLC tag table "250_TRANSP_PALLET_2"
   "_PALLET_EN_ALMACÉN" AT %M250.0 : Bool;
   "_PALLET_EN_ASCENSOR" AT %M250.1 : Bool;
   "_PALLET_EN_SEGURIDAD_ASCENS" AT %M250.2 : Bool;
   "_PALLET_EN_TRANSP_2" AT %M250.3 : Bool;
   "_PALLET_ENTRADA_ENVOLVEDORA" AT %M250.4 : Bool;
   "_PALLET_EN_ENVOLVEDORA" AT %M250.5 : Bool;
   "_PALLET_SALIDA_ENVOLVEDORA" AT %M250.6 : Bool;
   "_PALLET_EN_KETAN" AT %M250.7 : Bool;
   "_PALLET_EN_TRANSP_5" AT %M251.0 : Bool;
   "_PALLET_EN_DESCARGA" AT %M251.1 : Bool;
   "_Pedido_Recambio" AT %M251.2 : Bool;
   "_Retractilado" AT %M251.3 : Bool;
   "_Finciclo" AT %M251.4 : Bool;
END_VAR
